
   #sub_string := '';
   IF LEN(#str_in) >= #end_index AND #start_index < #end_index AND #start_index > 0 THEN
       #index := #start_index;
       WHILE #index <= #end_index DO
           #sub_string := CONCAT(IN1 := #sub_string, IN2 := #str_in[#index]);
           #index := #index + 1;
       END_WHILE;
   END_IF;
END_FUNCTION

FUNCTION "pa20b_station_monitoring" : Void   // FC59, SCL
{ S7_Optimized_Access := 'FALSE' }
VERSION : 0.1
BEGIN
   #pa20b_station_monitoring := false;
   IF #server_connection = true THEN

       IF #index = 255 THEN

               (* command *)
           Strg_TO_Chars(Strg := 'PA20B_STATE~',
                         pChars := 0,
                         Cnt => #chars,
                         Chars := #temp_buffer);
           #i := #chars;

           (* station state *)
           IF #station_activity_state = true THEN
               Strg_TO_Chars(Strg := 'Station state: Inactive~',
                             pChars := #i,
                             Cnt => #chars,
                             Chars := #temp_buffer);
           ELSE
               Strg_TO_Chars(Strg := 'Station state: Active~',
                             pChars := #i,
                             Cnt => #chars,
                             Chars := #temp_buffer);
           END_IF;

           #i := #i + #chars;

           (* cover release state *)
           IF #blend_senzor_l OR #blend_senzor_r THEN
               Strg_TO_Chars(Strg := 'Next cover expiration: Ready to remove~',
                             pChars := #i,
                             Cnt => #chars,
                             Chars := #temp_buffer);
           ELSE
               Strg_TO_Chars(Strg := 'Next cover expiration: Waiting~',
                             pChars := #i,
                             Cnt => #chars,
                             Chars := #temp_buffer);
           END_IF;

           #i := #i + #chars;
           #temp_buffer[#i] := '$L';

           #msg_index := "tcp_send"(#temp_buffer);
           IF #msg_index <> 255 THEN
               #index := #msg_index;
           END_IF;
       ELSE
           IF "tcp_rcv"(msg_index := #index, rcv_data => #temp_buffer) = true THEN
               #pa20b_station_monitoring := true;
               #index := 255;
           END_IF;
       END_IF;
   END_IF;
END_FUNCTION

FUNCTION "pa10b_station_monitoring" : Void   // FC60, SCL
{ S7_Optimized_Access := 'FALSE' }
VERSION : 0.1
BEGIN
   #pa10b_station_monitoring := false;
   IF #server_connection = true THEN

       IF #index = 255 THEN
       (* command *)
           Strg_TO_Chars(Strg := 'PA10B_STATE~',
                         pChars := 0,
                         Cnt => #chars,
                         Chars := #temp_buffer);
           #i := #chars;

           (* station state *)
           IF #station_activity_state = true THEN
               IF #fatal_error_state > 0 THEN
                   CASE #fatal_error_state OF
                       150:
                           Strg_TO_Chars(Strg := '<html>Station state: Y axis<br>valve lock error</html>~',
                                         pChars := #i,
                                         Cnt => #chars,
                                         Chars := #temp_buffer);
                       160:
                           Strg_TO_Chars(Strg := '<html>Station state: X axis<br>valve lock error</html>~',
                                         pChars := #i,
                                         Cnt => #chars,
                                         Chars := #temp_buffer);
                       ELSE
                           Strg_TO_Chars(Strg := 'Station state: Unknown~',
                                         pChars := #i,
                                         Cnt => #chars,
                                         Chars := #temp_buffer);
                   END_CASE;
               ELSE
                   IF #error_state > 0 THEN
                       Strg_TO_Chars(Strg := 'Station state: Unknown~',
                                     pChars := #i,
                                     Cnt => #chars,
                                     Chars := #temp_buffer);
                   ELSE
                       IF #big_fail_state > 0 THEN
                           CASE #big_fail_state OF
                               169:
                                   Strg_TO_Chars(Strg := 'Station state: Carring buffer inactive~',
                                                 pChars := #i,
                                                 Cnt => #chars,
                                                 Chars := #temp_buffer);
                               205:
                                   Strg_TO_Chars(Strg := 'Station state: Spacer in home position~',
                                                 pChars := #i,
                                                 Cnt => #chars,
                                                 Chars := #temp_buffer);
                               305:
                                   Strg_TO_Chars(Strg := 'Station state: Spacer out of home position~',
                                                 pChars := #i,
                                                 Cnt => #chars,
                                                 Chars := #temp_buffer);
                               ELSE  // Statement section ELSE
                                   Strg_TO_Chars(Strg := 'Station state: Unknown~',
                                                 pChars := #i,
                                                 Cnt => #chars,
                                                 Chars := #temp_buffer);
                           END_CASE;


                       ELSE
                           IF #fail_state > 0 THEN
                               CASE #fail_state OF
                                   150:
                                       Strg_TO_Chars(Strg := 'Station state: Felt box is empty~',
                                                     pChars := #i,
                                                     Cnt => #chars,
                                                     Chars := #temp_buffer);
                                   180:
                                       Strg_TO_Chars(Strg := 'Station state: Carring buffer inactive~',
                                                     pChars := #i,
                                                     Cnt => #chars,
                                                     Chars := #temp_buffer);
                                   203:
                                       Strg_TO_Chars(Strg := '<html>Station state: Activator bottle 1 in<br>primer box</html>~',
                                                     pChars := #i,
                                                     Cnt => #chars,
                                                     Chars := #temp_buffer);
                                   204:
                                       Strg_TO_Chars(Strg := '<html>Station state: Activator bottle 2 in<br>primer box</html>~',
                                                     pChars := #i,
                                                     Cnt => #chars,
                                                     Chars := #temp_buffer);
                                   205:
                                       Strg_TO_Chars(Strg := 'Station state: Spacer in home position~',
                                                     pChars := #i,
                                                     Cnt => #chars,
                                                     Chars := #temp_buffer);
                                   303:
                                       Strg_TO_Chars(Strg := '<html>Station state: Activator bottle 1<br>out of primer box</html>~',
                                                     pChars := #i,
                                                     Cnt => #chars,
                                                     Chars := #temp_buffer);
                                   304:
                                       Strg_TO_Chars(Strg := '<hrml>Station state: Activator bottle 2<br>out of primer box</html>~',
                                                     pChars := #i,
                                                     Cnt => #chars,
                                                     Chars := #temp_buffer);
                                   ELSE  // Statement section ELSE
                                       Strg_TO_Chars(Strg := 'Station state: Unknown~',
                                                     pChars := #i,
                                                     Cnt => #chars,
                                                     Chars := #temp_buffer);
                               END_CASE;

                           ELSE
                               Strg_TO_Chars(Strg := 'Station state: OK~',
                                             pChars := #i,
                                             Cnt => #chars,
                                             Chars := #temp_buffer);
                           END_IF;
                       END_IF;
                   END_IF;
               END_IF;
           ELSE
               Strg_TO_Chars(Strg := 'Station state: Inactive~',
                             pChars := #i,
                             Cnt => #chars,
                             Chars := #temp_buffer);
           END_IF;

           #i := #i + #chars;

           (* work cyclus state *)

           IF #work_cyclus_state = "RPA10B_hmi_go_to_home_position" THEN
               Strg_TO_Chars(Strg := 'Work cyclus state: Waiting for home position~',
                             pChars := #i,
                             Cnt => #chars,
                             Chars := #temp_buffer);
           ELSIF #work_cyclus_state = "RPA10B_hmi_scan_left_cover" THEN
               Strg_TO_Chars(Strg := 'Work cyclus state: Scan left cover code~',
                             pChars := #i,
                             Cnt => #chars,
                             Chars := #temp_buffer);
           ELSIF #work_cyclus_state = "RPA10B_hmi_scan_right_cover" THEN
               Strg_TO_Chars(Strg := 'Work cyclus state: Scan right cover code~',
                             pChars := #i,
                             Cnt => #chars,
                             Chars := #temp_buffer);
           ELSIF #work_cyclus_state = "RPA10B_hmi_move_roller_to_home_position" THEN
               Strg_TO_Chars(Strg := 'Work cyclus state: Move roller to home position~',
                             pChars := #i,
                             Cnt => #chars,
                             Chars := #temp_buffer);
           ELSIF #work_cyclus_state = "RPA10B_hmi_apply_activator_on_surface" THEN
               Strg_TO_Chars(Strg := '<html>Work cyclus state: Apply activator on surface and<br>put bottle back to primer box</html>~',
                             pChars := #i,
                             Cnt => #chars,
                             Chars := #temp_buffer);
           ELSIF #work_cyclus_state = "RPA10B_hmi_move_roller_to_left_cover" THEN
               Strg_TO_Chars(Strg := 'Work cyclus state: Mover roller to left cover~',
                             pChars := #i,
                             Cnt => #chars,
                             Chars := #temp_buffer);
           ELSIF #work_cyclus_state = "RPA10B_hmi_place_right_cover" THEN
               Strg_TO_Chars(Strg := 'Work cyclus state: Place right cover~',
                             pChars := #i,
                             Cnt => #chars,
                             Chars := #temp_buffer);
           ELSIF #work_cyclus_state = "RPA10B_hmi_place_left_cover" THEN
               Strg_TO_Chars(Strg := 'Work cyclus state: Place right cover~',
                             pChars := #i,
                             Cnt => #chars,
                             Chars := #temp_buffer);
           ELSIF #work_cyclus_state = "RPA10B_hmi_take_bottle_of_activator" THEN
               Strg_TO_Chars(Strg := 'Work cyclus state: Take bottle of activator~',
                             pChars := #i,
                             Cnt => #chars,
                             Chars := #temp_buffer);
           ELSIF #work_cyclus_state = "RPA10B_hmi_scan_bottle" THEN
               Strg_TO_Chars(Strg := 'Work cyclus state: Scan bottle of activator~',
                             pChars := #i,
                             Cnt => #chars,
                             Chars := #temp_buffer);
           ELSIF #work_cyclus_state = "RPA10B_hmi_change_pad" THEN
               Strg_TO_Chars(Strg := 'Work cyclus state: Change pad~',
                             pChars := #i,
                             Cnt => #chars,
                             Chars := #temp_buffer);
           ELSIF #work_cyclus_state = "RPA10B_hmi_apply_activator" THEN
               Strg_TO_Chars(Strg := 'Work cyclus state: Apply activator on cover surface~',
                             pChars := #i,
                             Cnt => #chars,
                             Chars := #temp_buffer);
           ELSIF #work_cyclus_state = "RPA10B_hmi_take_feld" THEN
               Strg_TO_Chars(Strg := 'Work cyclus state: Take felt from primer box~',
                             pChars := #i,
                             Cnt => #chars,
                             Chars := #temp_buffer);
           ELSIF #work_cyclus_state = "RPA10B_hmi_whipe_off" THEN
               Strg_TO_Chars(Strg := 'Work cyclus state: Whipe off~',
                             pChars := #i,
                             Cnt => #chars,
                             Chars := #temp_buffer);
           ELSIF #work_cyclus_state = "RPA10B_hmi_stick_sealing_on_right_cover" THEN
               Strg_TO_Chars(Strg := 'Work cyclus state: Stick sealing on right cover~',
                             pChars := #i,
                             Cnt => #chars,
                             Chars := #temp_buffer);
           ELSIF #work_cyclus_state = "RPA10B_hmi_press_universal_button_to_use_roller" THEN
               Strg_TO_Chars(Strg := '<html>Work cyclus state: Press universal button<br>to use roller</html>~',
                             pChars := #i,
                             Cnt => #chars,
                             Chars := #temp_buffer);
           ELSIF #work_cyclus_state = "RPA10B_hmi_Press_button_to_release_left_couver" THEN
               Strg_TO_Chars(Strg := '<html>Work cyclus state: Press button to<br>release left cover</html>~',
                             pChars := #i,
                             Cnt => #chars,
                             Chars := #temp_buffer);
           ELSIF #work_cyclus_state = "RPA10B_hmi_turn_fixture_to_left_cover" THEN
               Strg_TO_Chars(Strg := 'Work cyclus state: Turn fixture to left cover~',
                             pChars := #i,
                             Cnt => #chars,
                             Chars := #temp_buffer);
           ELSIF #work_cyclus_state = "RPA10B_hmi_turn_fixture_to_right_cover" THEN
               Strg_TO_Chars(Strg := 'Work cyclus state: Turn fixture to right cover~',
                             pChars := #i,
                             Cnt => #chars,
                             Chars := #temp_buffer);
           ELSIF #work_cyclus_state = "RPA10B_hmi_press_spacers_with_the_tool" THEN
               Strg_TO_Chars(Strg := 'Work cyclus state: Press spacer with the tool~',
                             pChars := #i,
                             Cnt => #chars,
                             Chars := #temp_buffer);
           ELSIF #work_cyclus_state = "RPA10B_hmi_press_button_to_release_right_couver" THEN
               Strg_TO_Chars(Strg := '<html>Work cyclus state: Press button to<br>release right cover</html>~',
                             pChars := #i,
                             Cnt => #chars,
                             Chars := #temp_buffer);
           ELSIF #work_cyclus_state = "RPA10B_cyclus_finished_OK" THEN
               Strg_TO_Chars(Strg := 'Work cyclus state: Work cyclus finished OK~',
                             pChars := #i,
                             Cnt => #chars,
                             Chars := #temp_buffer);
           ELSIF #work_cyclus_state = "RPA10B_hmi_active_carring_buffer" THEN
               Strg_TO_Chars(Strg := 'Work cyclus state: Active carring buffer~',
                             pChars := #i,
                             Cnt => #chars,
                             Chars := #temp_buffer);
           ELSIF #work_cyclus_state = "RPA10B_hmi_stick_sealing_on_left_cover" THEN
               Strg_TO_Chars(Strg := 'Work cyclus state: Stick sealing on left cover~',
                             pChars := #i,
                             Cnt => #chars,
                             Chars := #temp_buffer);
           ELSE
               Strg_TO_Chars(Strg := 'Work cyclus state: Unknown~',
                             pChars := #i,
                             Cnt => #chars,
                             Chars := #temp_buffer);
           END_IF;

           #i := #i + #chars;
           (* home position *)
           IF #position_sensor_2 AND #position_sensor_1 THEN
               Strg_TO_Chars(Strg := 'Home position: Yes~',
                             pChars := #i,
                             Cnt => #chars,
                             Chars := #temp_buffer);
           ELSE
               Strg_TO_Chars(Strg := 'Home position: No~',
                             pChars := #i,
                             Cnt => #chars,
                             Chars := #temp_buffer);
           END_IF;

           #i := #i + #chars;

           (* current left cover code *)
           Strg_TO_Chars(Strg := 'Current left cover code: ',
                         pChars := #i,
                         Cnt => #chars,
                         Chars := #temp_buffer);
           #i := #i + #chars;
           IF #current_left_cover_code <> '' THEN
               Strg_TO_Chars(Strg := #current_left_cover_code,
                             pChars := #i,
                             Cnt => #chars,
                             Chars := #temp_buffer);
           ELSE
               Strg_TO_Chars(Strg := 'None',
                             pChars := #i,
                             Cnt => #chars,
                             Chars := #temp_buffer);
           END_IF;
           #i := #i + #chars;

           (* current right cover code *)
           Strg_TO_Chars(Strg := '~Current right cover code: ',
                         pChars := #i,
                         Cnt => #chars,
                         Chars := #temp_buffer);
           #i := #i + #chars;

           IF #current_right_cover_code <> '' THEN
               Strg_TO_Chars(Strg := #current_right_cover_code,
                             pChars := #i,
                             Cnt => #chars,
                             Chars := #temp_buffer);
           ELSE
               Strg_TO_Chars(Strg := 'None',
                             pChars := #i,
                             Cnt => #chars,
                             Chars := #temp_buffer);
           END_IF;

           #i := #i + #chars;
           #temp_buffer[#i] := '$L';

           #msg_index := "tcp_send"(#temp_buffer);

           IF #msg_index <> 255 THEN
               #index := #msg_index;
           END_IF;
       ELSE
           IF "tcp_rcv"(msg_index := #index, rcv_data => #temp_buffer) = true THEN
               #pa10b_station_monitoring := true;
               #index := 255;
           END_IF;
       END_IF;
   END_IF;
END_FUNCTION

FUNCTION "tcp_send" : Void   // FC61, SCL
{ S7_Optimized_Access := 'FALSE' }
VERSION : 0.1
BEGIN
   (*
   send data on current buffer index to the pc, wait for the answare, the answare save to output buffer on the same index and 
   set the value in tcp_transaction_done on true
   *)


   IF (("tcp_datablock".index_out + 1) MOD 6) <> "tcp_datablock".index_send THEN
       IF "tcp_datablock".tcp_transaction_done["tcp_datablock".index_out] = false THEN
           WHILE #data[#index] <> '$L' DO
               "tcp_datablock".tcp_output_buffer["tcp_datablock".index_out].tcp_item[#index] := #data[#index];
               #index := #index + 1;
           END_WHILE;

           "tcp_datablock".tcp_size_out["tcp_datablock".index_out] := #index;
           #tcp_send := "tcp_datablock".index_out;

       ELSE
           #tcp_send := 255;
       END_IF;
       "tcp_datablock".index_out := ("tcp_datablock".index_out +1) MOD 6;
   ELSE
       #tcp_send := 255;
   END_IF;
END_FUNCTION

FUNCTION "RPA20B_handler_op_1" : Void   // FC62, SCL
{ S7_Optimized_Access := 'FALSE' }
VERSION : 0.1
BEGIN
   "RPA20_motor_up" := false;

   IF "RPA20B_ES_feedback" = false THEN

       "IEC_Timer_0_DB".TON(IN := "RPA20B_Camera_Start_Test",
                            PT := T#200ms);

       IF "RPA20B_Camera_Start_Test" AND "IEC_Timer_0_DB".Q AND ("RPA20B_Camera_Test_Ok"=TRUE OR "RPA20B_Product_Present_On_Top_Level"=FALSE) THEN
           "RPA20B_Camera_Result_OK" := TRUE;
           "RPA20B_Camera_Result_NOK" := FALSE;
       END_IF;
       IF "RPA20B_Camera_Start_Test" AND "IEC_Timer_0_DB".Q AND "RPA20B_Camera_Test_Ok" = FALSE AND "RPA20B_Product_Present_On_Top_Level" = TRUE THEN
           "RPA20B_Camera_Result_OK" := FALSE;
           "RPA20B_Camera_Result_NOK" := TRUE;
       END_IF;

       "PA20B_Timer_0_DB".TON(IN := "RPA20B_Camera_Result_OK",
                              PT := T#2m);

       IF "RPA20B_Camera_Result_OK" = TRUE THEN
           IF "PA20B_Timer_0_DB".Q = true THEN
               "RPA20B_datablock".RPA20B_buffer_down_enable := true;
               "RPA20B_Camera_Result_OK" := FALSE;
               "RPA20B_Camera_Result_NOK" := FALSE;
           END_IF;

       END_IF;

       IF "RPA20B_datablock".RPA20B_automatic_cyclus_enable = true THEN
       (* main cyclus *)
           CASE "RPA20B_datablock".RPA20B_work_cyclus_state_OP_1 OF
               0: // init
                   "RPA20B_motor_down" := NOT "RPA20B_belt_position_sensor" AND (NOT "RPA20B_open_drawer");
                   IF "RPA20B_belt_position_sensor" = true THEN
                       "RPA20B_datablock".RPA20B_work_cyclus_state_OP_1 := 1;
                   END_IF;
               1:
                   IF ("RPA20B_blend_presence_sensor_1" = false AND "RPA20B_blend_presence_sensor_2" = false) THEN
                       IF "RPA20B_datablock".RPA20B_buffer_down_enable = true THEN
                           "RPA20B_datablock".RPA20B_buffer_down_enable := false;
                           "RPA20B_datablock".RPA20B_work_cyclus_state_OP_1 := 3;
                       END_IF;
                   ELSE
                       "RPA20B_datablock".RPA20B_automatic_cyclus_enable := false;
                   END_IF;
               3:
                   "RPA20B_motor_down" := true;
                   IF "RPA20B_belt_position_sensor" = false THEN
                       "RPA20B_datablock".RPA20B_work_cyclus_state_OP_1 := 4;
                   END_IF;
               4:
                   "RPA20B_motor_down" := true;
                   IF "RPA20B_belt_position_sensor" = true THEN
                       "RPA20B_datablock".RPA20B_work_cyclus_state_OP_1 := 0;
                       "RPA20B_motor_down" := false;
                   END_IF;
               ELSE
                   "RPA20B_datablock".RPA20B_work_cyclus_state_OP_1 := 0;
                   "RPA20B_datablock".RPA20B_buffer_down_enable := false;
                   "RPA20B_motor_down" := false;
           END_CASE;
       ELSE
           IF "RPA20B_open_drawer" = false AND "PA20B_Timer_1_DB".Q = true THEN
               "RPA20B_datablock".RPA20B_automatic_cyclus_enable := true;
           ELSE
               "RPA20B_motor_down" := false;
               "RPA20B_datablock".RPA20B_automatic_cyclus_enable := false;
           END_IF;

           "PA20B_Timer_1_DB".TON(IN := ("RPA20B_open_drawer" = false AND ("RPA20B_blend_presence_sensor_1" = false AND "RPA20B_blend_presence_sensor_2" = false)),
                                  PT := T#10s);
       END_IF;

       (* cover demage protection *)
       IF "RPA20B_open_drawer" = true THEN
           "RPA20B_datablock".RPA20B_automatic_cyclus_enable := false;
       END_IF;
   END_IF;
END_FUNCTION

FUNCTION "RPA10B_change_pad" : Void   // FC63, SCL
{ S7_Optimized_Access := 'FALSE' }
VERSION : 0.1
BEGIN



   IF "checkFailStateLock"(failStateLock := #failStatelockIdetifier,
                                       bigFailStateLock := #bigFailStateLock,
                                       ErrorStateLock := #bigFailStateLock,
                                       FatalErrorStateLock := #FatalErrorStateLock,
                                       failStatelockIdetifier := #failStatelockIdetifier) THEN

       #readyLED := (NOT  "RPA10B_datablock".RPA10B_pad_checking_trigr) AND #padIsChangedButton;
       #notReadyLED := NOT #readyLED;

       #RPA10B_change_pad := #readyLED;

       IF #padSensor = false AND "RPA10B_datablock".RPA10B_pad_checking_trigr = true THEN
           #changePedLED := "Clock_0.5Hz";
           IF #padIsChangedButton THEN
               #RPA10B_change_pad := true;
               "setOKState"(confirm := true,
                            identifier := #failStatelockIdetifier,
                            confirm_blinking := false,
                            blinkConfirmButton => #confirmButtonLED,
                            stateLock := #failStateLock);
               "RPA10B_datablock".RPA10B_pad_checking_trigr := false;
               #changePedLED := false;
           END_IF;
       ELSE
           #changePedLED := #notReadyLED;
           #RPA10B_change_pad := false;
           IF "setFailState"(identifier := #failStatelockIdetifier,
                                 failStateLock := #failStateLock) THEN
               ;
           END_IF;
       END_IF;

       "RPA10B_datablock".RPA10B_pad_checking_trigr := #padSensor OR "RPA10B_datablock".RPA10B_pad_checking_trigr;
   ELSE
       #RPA10B_change_pad := false;
   END_IF;
END_FUNCTION

FUNCTION "RPA20B_handler_op_2" : Void   // FC64, SCL
{ S7_Optimized_Access := 'FALSE' }
VERSION : 0.1
BEGIN
   CASE "RPA20B_datablock".RPA20B_work_cyclus_state_OP_2 OF

       "RPA20B_blend_expiration_checking":
           IF "RPA20B_blend_presence_sensor_1" = true OR "RPA20B_blend_presence_sensor_2" = true AND "RPA20B_motor_down" = false THEN
               "RPA20B_datablock".RPA20B_work_cyclus_state_OP_2 := "RPA20B_wait_to_push_open_button";
           ELSE
               "RPA20B_valve_close_drawer" := true;
               "RPA20B_valve_open_drawer" := false;
               "RPA20B_open_drawer" := false;
           END_IF;

       "RPA20B_wait_to_push_open_button":
               IF "RPA20B_unlock_button" = true AND "RPA20B_motor_down" = false THEN
                   IF "RPA20B_blend_presence_sensor_1" = true OR "RPA20B_blend_presence_sensor_2" = true THEN
                       "RPA20B_valve_close_drawer" := false;
                       "RPA20B_valve_open_drawer" := true;
                       "RPA20B_open_drawer" := true;
                       "RPA20B_datablock".RPA20B_work_cyclus_state_OP_2 := "RPA20B_wait_for_deactivate_open_button";
                   ELSE
                       "RPA20B_datablock".RPA20B_work_cyclus_state_OP_2 := "RPA20B_blend_expiration_checking";
                   END_IF;
               END_IF;

       "RPA20B_wait_for_deactivate_open_button":
           IF "RPA20B_unlock_button" = false THEN
               "RPA20B_datablock".RPA20B_work_cyclus_state_OP_2 := "RPA20B_wait_to_push_close_button";
           END_IF;

       "RPA20B_wait_to_push_close_button":
           IF "RPA20B_unlock_button" = true AND "RPA20B_drawer_lock_sensor" = false AND "RPA20B_drawer_position_sensor" = true AND "RPA20B_drawer_unlock_sensor" = true THEN
               "RPA20B_valve_close_drawer" := true;
               "RPA20B_valve_open_drawer" := false;
               "RPA20B_datablock".RPA20B_work_cyclus_state_OP_2 := "RPA20B_is_blend_release";
           END_IF;

       "RPA20B_is_blend_release":
           IF "RPA20B_drawer_lock_sensor" = true AND "RPA20B_drawer_unlock_sensor" = false THEN
               IF "RPA20B_blend_presence_sensor_1" = false AND "RPA20B_blend_presence_sensor_2" = false THEN
                   "RPA20B_datablock".RPA20B_work_cyclus_state_OP_2 := "RPA20B_end_operation";
                   "RPA20B_open_drawer" := false;
               ELSE
                   "RPA20B_valve_close_drawer" := false;
                   "RPA20B_valve_open_drawer" := true;
                   "RPA20B_datablock".RPA20B_work_cyclus_state_OP_2 := "RPA20B_wait_for_deactivate_open_button";
               END_IF;
           END_IF;

       "RPA20B_end_operation":
           IF "RPA20B_unlock_button" = false THEN
               "RPA20B_datablock".RPA20B_work_cyclus_state_OP_2 := "RPA20B_blend_expiration_checking";
           END_IF;

       ELSE  // Statement section ELSE
           "RPA20B_datablock".RPA20B_work_cyclus_state_OP_2 := "RPA20B_blend_expiration_checking";
           "RPA20B_valve_close_drawer" := true;
           "RPA20B_valve_open_drawer" := false;
           "RPA20B_open_drawer" := false;
   END_CASE;
END_FUNCTION

FUNCTION "tcp_rcv" : Void   // FC65, SCL
{ S7_Optimized_Access := 'FALSE' }
VERSION : 0.1
BEGIN
   (*

   *)

   #tcp_rcv := false;

   IF "tcp_datablock".tcp_transaction_done[#msg_index] = true THEN
       WHILE #index < 1023 DO
           #rcv_data[#index] := "tcp_datablock".tcp_input_buffer[#msg_index].tcp_item[#index];
           #index := #index + 1;
       END_WHILE;
       "tcp_datablock".tcp_transaction_done[#msg_index] := false;
       #tcp_rcv := true;
   END_IF;
END_FUNCTION

FUNCTION "tcp_runtime" : Void   // FC66, SCL
{ S7_Optimized_Access := 'FALSE' }
VERSION : 0.1
BEGIN
   (*

   *)


   IF "tcp_datablock".tcp_connection = true THEN
       IF "tcp_datablock".index_send <> "tcp_datablock".index_out THEN
           IF "tcp_datablock"."counter" > 0 THEN
               "tcp_datablock"."counter" := "tcp_datablock"."counter" - 1;
               IF "tcp_datablock".tcp_transaction_done["tcp_datablock".index_send] = false THEN
                   IF "TCP_TSEND_DB".DONE = false THEN
                       "TCP_TSEND_DB".REQ := NOT "TCP_TSEND_DB".REQ;
                       "tcp_datablock".tcp_output_buffer["tcp_datablock".index_send].tcp_item["tcp_datablock".tcp_size_out["tcp_datablock".index_send]] := '$R';
                        "tcp_datablock".tcp_output_buffer["tcp_datablock".index_send].tcp_item["tcp_datablock".tcp_size_out["tcp_datablock".index_send]+1] := '$L';

                        "TCP_TSEND_DB".TSEND(DATA := "tcp_datablock".tcp_output_buffer["tcp_datablock".index_send].tcp_item,
                                                LEN := "tcp_datablock".tcp_size_out["tcp_datablock".index_send]+2,
                                                ID := 2);
                   ELSE
                       IF "TCP_TRCV_DB".NDR = false THEN
                           "TCP_TRCV_DB".TRCV(EN_R := true,
                                              ID := 2,
                                              LEN := 1024,
                                              DATA := "tcp_datablock".tcp_input_buffer["tcp_datablock".index_send].tcp_item);
                       ELSE
                           "tcp_datablock"."counter" := 1024;
                           "TCP_TRCV_DB".NDR := false;
                           "TCP_TSEND_DB".DONE := false;
                           "tcp_datablock".tcp_transaction_done["tcp_datablock".index_send] := true;
                           "tcp_datablock".index_send := ("tcp_datablock".index_send + 1) MOD 6;
                       END_IF;
                   END_IF;
               ELSE
                   "tcp_datablock".index_send := ("tcp_datablock".index_send + 1) MOD 6;
               END_IF;
           ELSE
               "TCP_TRCV_DB".NDR := false;
               "TCP_TSEND_DB".DONE := false;
               "tcp_datablock".tcp_connection := false;
           END_IF;
       END_IF;
   ELSE
       "TCP_TRCV_DB".NDR := false;
       "TCP_TSEND_DB".DONE := false;
   END_IF;
END_FUNCTION

FUNCTION "tcp_connect" : Void   // FC67, SCL
{ S7_Optimized_Access := 'FALSE' }
VERSION : 0.1
BEGIN
   (*

   *)

   IF "tcp_datablock".tcp_connection = false THEN
       IF "tcp_datablock"."counter" > 0 THEN
           "tcp_datablock"."counter" := "tcp_datablock"."counter" - 1;

           IF "TCP_TDISCON_DB".DONE = false AND "TCP_TDISCON_DB".STATUS <> 16#80A3 THEN
               "TCP_TDISCON_DB".REQ := (NOT "TCP_TDISCON_DB".REQ);
               "TCP_TDISCON_DB"(ID := 2);
           ELSE
               IF "TCP_TCON_DB".DONE = false THEN
                   "TCP_TCON_DB".REQ := NOT "TCP_TCON_DB".REQ;
                   "TCP_TCON_DB"(CONNECT := "TCP_Connection_DB",
                                  ID := 2);
               ELSE
                   "tcp_datablock".tcp_connection := true;
                   "tcp_datablock"."counter" := 1024;
                   "TCP_TCON_DB".DONE := false;
                   "TCP_TDISCON_DB".DONE := false;
                   "TCP_TDISCON_DB".STATUS := 0;
               END_IF;
           END_IF;
       ELSE
           "tcp_datablock"."counter" := 1024;
           "TCP_TCON_DB".DONE := false;
           "TCP_TDISCON_DB".DONE := false;
           "TCP_TDISCON_DB".STATUS := 0;
       END_IF;
   END_IF;
END_FUNCTION

FUNCTION "generate_csv" : Void   // FC69, SCL
{ S7_Optimized_Access := 'FALSE' }
VERSION : 0.1
BEGIN
   #generate_csv := false;

   IF #server_conection = true THEN
       IF #index = 255 THEN

           #temp_string := CONCAT(IN1 :='GENERATE_CSV~' , IN2 :=#record );

           IF #frame = 0 THEN
               #temp_string := CONCAT(IN1 := #temp_string, IN2 := '~glued_frame_581~0~0$L');
           ELSE
               #temp_string := CONCAT(IN1 := #temp_string, IN2 := '~glued_frame_AU326_1~0~0$L');
           END_IF;

           Strg_TO_Chars(Strg := #temp_string,
                         pChars := 0,
                         Cnt => #chars,
                         Chars := #record_buffer);

           #msg_index := "tcp_send"(#record_buffer);

           IF #msg_index <> 255 THEN
               #index := #msg_index;
           END_IF;
       ELSE
           IF "tcp_rcv"(msg_index := #index, rcv_data => #record_buffer) = true THEN
               #generate_csv := true;
               #index := 255;
           END_IF;
       END_IF;
   END_IF;
END_FUNCTION

FUNCTION "parse_scanned_label" : Void   // FC70, SCL
{ S7_Optimized_Access := 'FALSE' }
VERSION : 0.1
BEGIN

   IF #scanned_data[LEN(#scanned_data)] = 'M' OR #scanned_data[LEN(#scanned_data)] = 'S' THEN

       #index := 1;
       WHILE #scanned_data[#index] <> '*' AND #index < LEN(#scanned_data) DO
           #chemical := CONCAT(IN1 := #chemical, IN2 := #scanned_data[#index]);
           #index := #index + 1;
       END_WHILE;

       (* batch code *)
       #index := #index + 1;
       WHILE #scanned_data[#index] <> '*' AND #index < LEN(#scanned_data) DO
           #batch_no := CONCAT(IN1 := #batch_no, IN2 := #scanned_data[#index]);
           #index := #index + 1;
       END_WHILE;

       #expire_date_time.DAY := STRING_TO_USINT("sub_string"(str_in := #scanned_data, start_index := #index + 1, end_index := #index + 2));
       #expire_date_time.MONTH := STRING_TO_USINT("sub_string"(str_in := #scanned_data, start_index := #index + 4, end_index := #index + 5));
       #expire_date_time.YEAR := STRING_TO_UINT("sub_string"(str_in := #scanned_data, start_index := #index + 7, end_index := #index + 10));
       #expire_date_time.HOUR := STRING_TO_USINT("sub_string"(str_in := #scanned_data, start_index := #index + 12, end_index := #index + 13));
       #expire_date_time.MINUTE := STRING_TO_USINT("sub_string"(str_in := #scanned_data, start_index := #index + 15, end_index := #index + 16));

       #index := #index + 17;

       #filling_opening_date_time.DAY := STRING_TO_USINT("sub_string"(str_in := #scanned_data, start_index := #index + 1, end_index := #index + 2));
       #filling_opening_date_time.MONTH := STRING_TO_USINT("sub_string"(str_in := #scanned_data, start_index := #index + 4, end_index := #index + 5));
       #filling_opening_date_time.YEAR := STRING_TO_UINT("sub_string"(str_in := #scanned_data, start_index := #index + 7, end_index := #index + 10));
       #filling_opening_date_time.HOUR := STRING_TO_USINT("sub_string"(str_in := #scanned_data, start_index := #index + 12, end_index := #index + 13));
       #filling_opening_date_time.MINUTE := STRING_TO_USINT("sub_string"(str_in := #scanned_data, start_index := #index + 15, end_index := #index + 16));

       #index := #index + 1;
       (* opening date *)
       WHILE #scanned_data[#index] <> '*' AND #index < LEN(#scanned_data) DO
           #index := #index + 1;
       END_WHILE;

       (* opening time *)
       #index := #index + 1;
       WHILE #scanned_data[#index] <> '*' AND #index < LEN(#scanned_data) DO
           #index := #index + 1;
       END_WHILE;

       #bottle_type := #scanned_data[LEN(#scanned_data)];
   ELSE
       #bottle_type := 'U';
   END_IF;
END_FUNCTION

FUNCTION "fs_internal_state" : Void   // FC71, SCL
{ S7_Optimized_Access := 'FALSE' }
VERSION : 0.1
BEGIN
   IF #switch_automat_manual = true THEN
       #error_state := 2;
   END_IF;

   IF #switch_automat_manual = false AND #error_state = 2 THEN
       #error_state := 0;
   END_IF;

   IF #tcp_connection = false THEN
       #error_state := 1;
   END_IF;

   IF #tcp_connection = true AND #error_state = 1 THEN
       #error_state := 0;
   END_IF;

   (* error state reset *)
   IF #confirm_button = true THEN
       #error_state := 0;
   END_IF;

   (* beacon and siren *)
   IF #error_state = 0 THEN
       #beacon_green := true;
       #beacon_red := false;
       #beacon_orange := false;
       #alarm := false;
   ELSE
       #beacon_green := false;
       #beacon_red := true;
       #beacon_orange := false;
       #alarm := true;
   END_IF;

   IF #error_state > 255 THEN
       #beacon_siren := true;
   ELSE
       #beacon_siren := false;
   END_IF;

   #confirm_led := #beacon_red;
END_FUNCTION

FUNCTION "station_inactive_state" : Void   // FC72, SCL
{ S7_Optimized_Access := 'FALSE' }
VERSION : 0.1
BEGIN


   "station_reset"(funel_1:=#fune_1,
                   funel_2:=#fune_2,
                   funel_3:=#fune_3,
                   funel_4:=#fune_4,
                   funel_5:=#fune_5,
                   fs_reset_e:=#fs_reset_enable,
                   fs_chemical_type:=#chemical_type,
                   fill_bottle_step:=#fill_bottle_step,
                   shake_deinit:=#shake_deinit,
                   print_sp_bottle_label_step:=#print_sp_bottle_label_step,
                   fs_show_manual_or_scan:=#fs_show_manual_or_scan,
                   fs_show_button:=#fs_show_button,
                   fs_show_fill_button:=#fs_show_fill_button,
                   fs_funel_control:=#fs_funel_control,
                   hmi_label_index:=#hmi_label_index);
   #error_state := 0;
   #beacon_red := false;
   #beacon_green := false;
   #beacon_orange := false;
   #beacon_siren := false;

   #fs_start_led := "Clock_0.5Hz";
   IF #fs_start_button = true THEN
       #fs_station_activity := true;
       #fs_start_led := false;
   END_IF;
END_FUNCTION

ORGANIZATION_BLOCK "Main"   // OB1, LAD, ProgramCycle
TITLE = "Main Program Sweep (Cycle)"
{ S7_Optimized_Access := 'FALSE' }
VERSION : 0.1
BEGIN

REGION Network 1
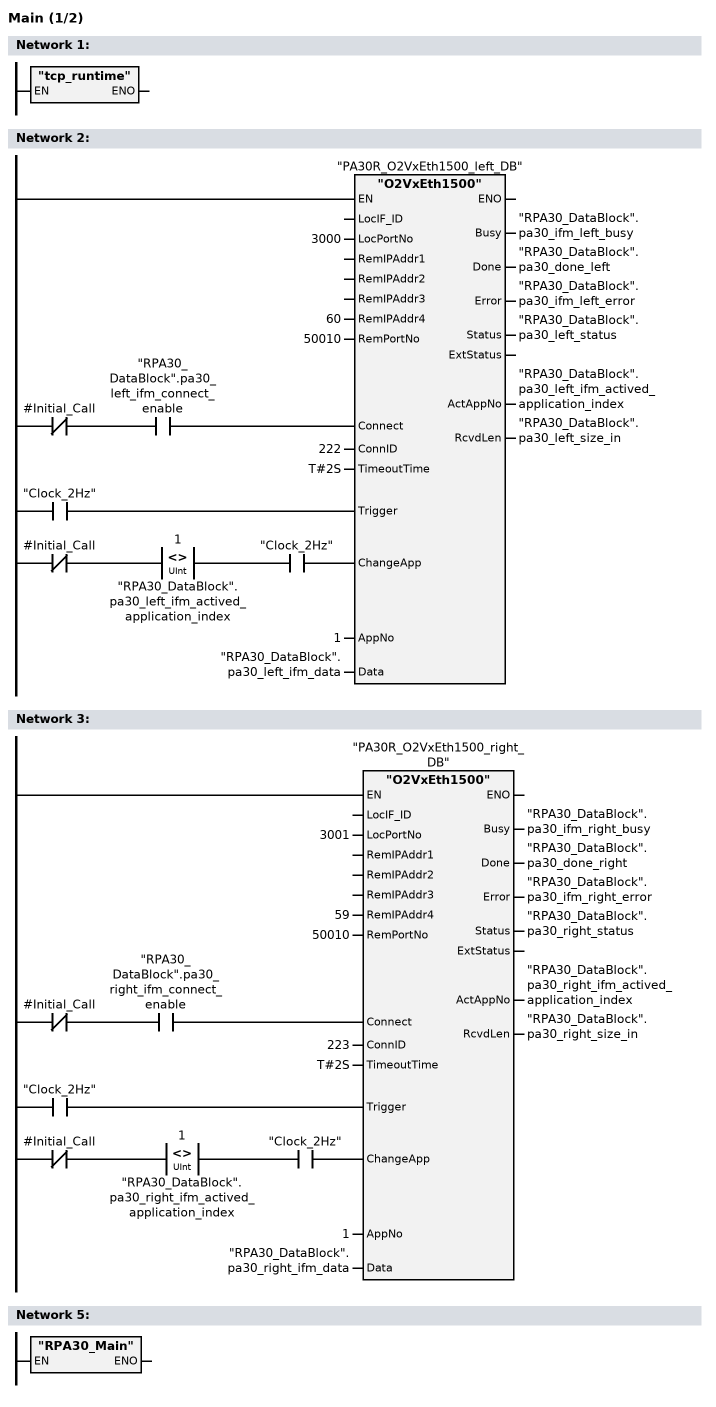
   RUNG wire#powerrail
      "tcp_runtime"()
   END_RUNG
   // the same network as SCL:
   "tcp_runtime"();
END_REGION

REGION Network 2
   RUNG wire#powerrail
      "PA30R_O2VxEth1500_left_DB"(Connect := wire#w1, Trigger := wire#w2, ChangeApp := wire#w3, LocIF_ID :=, LocPortNo := 3000, RemIPAddr1 :=, RemIPAddr2 :=, RemIPAddr3 :=, RemIPAddr4 := 60, RemPortNo := 50010, ConnID := 222, TimeoutTime := T#2S, AppNo := 1, Data := "RPA30_DataBlock".pa30_left_ifm_data, Busy => "RPA30_DataBlock".pa30_ifm_left_busy, Done => "RPA30_DataBlock".pa30_done_left, Error => "RPA30_DataBlock".pa30_ifm_left_error, Status => "RPA30_DataBlock".pa30_left_status, ExtStatus =>, ActAppNo => "RPA30_DataBlock".pa30_left_ifm_actived_application_index, RcvdLen => "RPA30_DataBlock".pa30_left_size_in)
   END_RUNG
   RUNG wire#powerrail
      I_Contact( #Initial_Call )
      Contact( "RPA30_DataBlock".pa30_left_ifm_connect_enable )
   END_RUNG wire#w1
   RUNG wire#powerrail
      Contact( "Clock_2Hz" )
   END_RUNG wire#w2
   RUNG wire#powerrail
      I_Contact( #Initial_Call )
      { S7_Templates := "SrcType := UInt" } NE_Contact(in1 := 1, in2 := "RPA30_DataBlock".pa30_left_ifm_actived_application_index)
      Contact( "Clock_2Hz" )
   END_RUNG wire#w3
   // the same network as SCL:
   "PA30R_O2VxEth1500_left_DB"(LocPortNo := 3000,   // "O2VxEth1500"
                           RemIPAddr4 := 60,
                           RemPortNo := 50010,
                           Connect := NOT #Initial_Call AND "RPA30_DataBlock".pa30_left_ifm_connect_enable,
                           ConnID := 222,
                           TimeoutTime := T#2S,
                           Trigger := "Clock_2Hz",
                           ChangeApp := NOT #Initial_Call AND (1 <> "RPA30_DataBlock".pa30_left_ifm_actived_application_index) AND "Clock_2Hz",
                           AppNo := 1,
                           Data := "RPA30_DataBlock".pa30_left_ifm_data,
                           Busy => "RPA30_DataBlock".pa30_ifm_left_busy,
                           Done => "RPA30_DataBlock".pa30_done_left,
                           Error => "RPA30_DataBlock".pa30_ifm_left_error,
                           Status => "RPA30_DataBlock".pa30_left_status,
                           ActAppNo => "RPA30_DataBlock".pa30_left_ifm_actived_application_index,
                           RcvdLen => "RPA30_DataBlock".pa30_left_size_in);
END_REGION

REGION Network 3
   RUNG wire#powerrail
      "PA30R_O2VxEth1500_right_DB"(Connect := wire#w1, Trigger := wire#w2, ChangeApp := wire#w3, LocIF_ID :=, LocPortNo := 3001, RemIPAddr1 :=, RemIPAddr2 :=, RemIPAddr3 :=, RemIPAddr4 := 59, RemPortNo := 50010, ConnID := 223, TimeoutTime := T#2S, AppNo := 1, Data := "RPA30_DataBlock".pa30_right_ifm_data, Busy => "RPA30_DataBlock".pa30_ifm_right_busy, Done => "RPA30_DataBlock".pa30_done_right, Error => "RPA30_DataBlock".pa30_ifm_right_error, Status => "RPA30_DataBlock".pa30_right_status, ExtStatus =>, ActAppNo => "RPA30_DataBlock".pa30_right_ifm_actived_application_index, RcvdLen => "RPA30_DataBlock".pa30_right_size_in)
   END_RUNG
   RUNG wire#powerrail
      I_Contact( #Initial_Call )
      Contact( "RPA30_DataBlock".pa30_right_ifm_connect_enable )
   END_RUNG wire#w1
   RUNG wire#powerrail
      Contact( "Clock_2Hz" )
   END_RUNG wire#w2
   RUNG wire#powerrail
      I_Contact( #Initial_Call )
      { S7_Templates := "SrcType := UInt" } NE_Contact(in1 := 1, in2 := "RPA30_DataBlock".pa30_right_ifm_actived_application_index)
      Contact( "Clock_2Hz" )
   END_RUNG wire#w3
   // the same network as SCL:
   "PA30R_O2VxEth1500_right_DB"(LocPortNo := 3001,   // "O2VxEth1500"
                           RemIPAddr4 := 59,
                           RemPortNo := 50010,
                           Connect := NOT #Initial_Call AND "RPA30_DataBlock".pa30_right_ifm_connect_enable,
                           ConnID := 223,
                           TimeoutTime := T#2S,
                           Trigger := "Clock_2Hz",
                           ChangeApp := NOT #Initial_Call AND (1 <> "RPA30_DataBlock".pa30_right_ifm_actived_application_index) AND "Clock_2Hz",
                           AppNo := 1,
                           Data := "RPA30_DataBlock".pa30_right_ifm_data,
                           Busy => "RPA30_DataBlock".pa30_ifm_right_busy,
                           Done => "RPA30_DataBlock".pa30_done_right,
                           Error => "RPA30_DataBlock".pa30_ifm_right_error,
                           Status => "RPA30_DataBlock".pa30_right_status,
                           ActAppNo => "RPA30_DataBlock".pa30_right_ifm_actived_application_index,
                           RcvdLen => "RPA30_DataBlock".pa30_right_size_in);
END_REGION

REGION Network 5
   RUNG wire#powerrail
      "RPA30_Main"()
   END_RUNG
   // the same network as SCL:
   "RPA30_Main"();
END_REGION

REGION Network 7
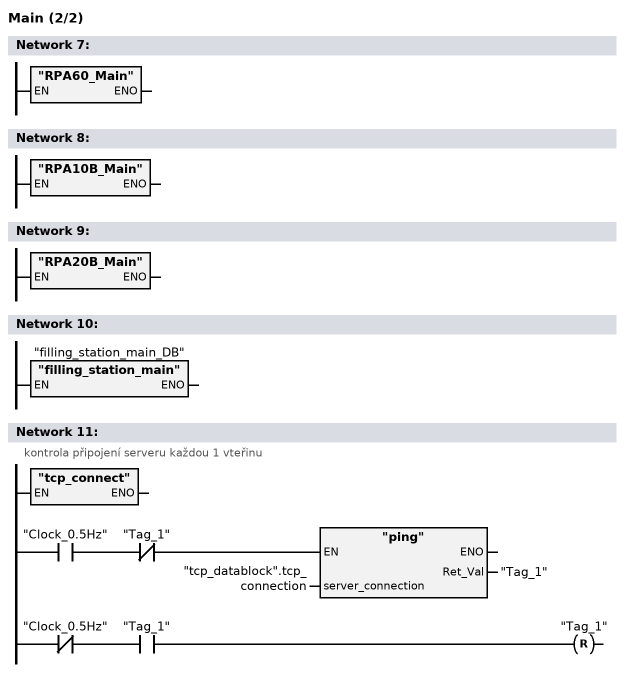
   RUNG wire#powerrail
      "RPA60_Main"()
   END_RUNG
   // the same network as SCL:
   "RPA60_Main"();
END_REGION

REGION Network 8
   RUNG wire#powerrail
      "RPA10B_Main"()
   END_RUNG
   // the same network as SCL:
   "RPA10B_Main"();
END_REGION

REGION Network 9
   RUNG wire#powerrail
      "RPA20B_Main"()
   END_RUNG
   // the same network as SCL:
   "RPA20B_Main"();
END_REGION

REGION Network 10
   RUNG wire#powerrail
      "filling_station_main_DB"()
   END_RUNG
   // the same network as SCL:
   "filling_station_main_DB"();   // "filling_station_main"
END_REGION

REGION Network 11
   // kontrola připojení serveru každou 1 vteřinu
   RUNG wire#powerrail
      "tcp_connect"()
   END_RUNG
   RUNG wire#powerrail
      Contact( "Clock_0.5Hz" )
      I_Contact( "Tag_1" )
      "ping"(server_connection := "tcp_datablock".tcp_connection, Ret_Val => "Tag_1")
   END_RUNG
   RUNG wire#powerrail
      I_Contact( "Clock_0.5Hz" )
      Contact( "Tag_1" )
      R_Coil( "Tag_1" )
   END_RUNG
   // the same network as SCL:
   "tcp_connect"();
   IF "Clock_0.5Hz" AND NOT "Tag_1" THEN
       "Tag_1" := "ping"(server_connection := "tcp_datablock".tcp_connection);
   END_IF;
   IF NOT "Clock_0.5Hz" AND "Tag_1" THEN "Tag_1" := FALSE; END_IF;
END_REGION
END_ORGANIZATION_BLOCK

ORGANIZATION_BLOCK "CyclicInterrupt_Ms"   // OB32, SCL, CyclicInterrupt
{ S7_Optimized_Access := 'FALSE' }
VERSION : 0.1
BEGIN

   IF NOT "RPA30R_LCDSwitchAutomat_Manual" THEN
       IF "RPA30_DataBlock".RPA30_valveYErrorStateCheck > 0 THEN

           "RPA30_DataBlock".RPA30_valveYErrorStateCheck := "RPA30_DataBlock".RPA30_valveYErrorStateCheck - 1;
       END_IF;

       IF "RPA60_DataBlock".RPA60_valveYErrorStateCheck > 0 THEN

           "RPA60_DataBlock".RPA60_valveYErrorStateCheck := "RPA60_DataBlock".RPA60_valveYErrorStateCheck - 1;
       END_IF;
   END_IF;

   IF "RPA10B_datablock".RPA10B_vacuum_R_check_state > 0 THEN
       "RPA10B_datablock".RPA10B_vacuum_R_check_state :="RPA10B_datablock".RPA10B_vacuum_R_check_state - 1;
   END_IF;

   IF "RPA10B_datablock".RPA10B_vacuum_L_check_state > 0 THEN
       "RPA10B_datablock".RPA10B_vacuum_L_check_state := "RPA10B_datablock".RPA10B_vacuum_L_check_state - 1;
   END_IF;

   IF "RPA10B_datablock".RPA10_valve_Y_check_state > 0 THEN
       "RPA10B_datablock".RPA10_valve_Y_check_state := "RPA10B_datablock".RPA10_valve_Y_check_state - 1;
   END_IF;

   IF "RPA10B_datablock".RPA10_valve_X_check_state > 0 THEN
       "RPA10B_datablock".RPA10_valve_X_check_state := "RPA10B_datablock".RPA10_valve_X_check_state - 1;
   END_IF;
END_ORGANIZATION_BLOCK

(* ===== HMI "HMI_RT_2" =====
connection "HMI_Connection_2": ETHERNET, SMART_S7_1500_OMS

